   286: 'IGG_MESSAGE_WORD_02_BIT_5', class IGG Messages, trigger "64_Message_Data_IGG_MESSAGE_WORD_02" bit 13
   126: 'PIT-113 IGG MAIN ATOM AIR PRESSURE - FAULT', class BC Alarms, trigger "BC_ALARM_ACKNLG_4" bit 13
   125: 'TS-403 IG TEMP - HIGH HIGH SWITCH AND TIT-360 - FAULT', class BC Alarms, trigger "BC_ALARM_ACKNLG_4" bit 12
   128: 'TIT-202 IGG INLET FUEL TEMP', class BC Alarms, trigger "BC_ALARM_ACKNLG_4" bit 15
   127: 'PIT-205 IGG MAIN FUEL PRESSURE - FAULT', class BC Alarms, trigger "BC_ALARM_ACKNLG_4" bit 14
   313: 'BC_MESSAGE_WORD_02_BIT_0', class BC Messages, trigger "64_Message_Data_BC_MESSAGE_WORD_02" bit 8
   292: 'BC_MESSAGE_WORD_01_BIT_11', class BC Messages, trigger "64_Message_Data_BC_MESSAGE_WORD_01" bit 3
   311: 'BC_MESSAGE_WORD_02_BIT_14', class BC Messages, trigger "64_Message_Data_BC_MESSAGE_WORD_02" bit 6
   312: 'BC_MESSAGE_WORD_02_BIT_15', class BC Messages, trigger "64_Message_Data_BC_MESSAGE_WORD_02" bit 7
   289: 'BC_MESSAGE_WORD_01_BIT_8', class BC Messages, trigger "64_Message_Data_BC_MESSAGE_WORD_01" bit 0
   288: 'IGG_MESSAGE_WORD_02_BIT_7', class IGG Messages, trigger "64_Message_Data_IGG_MESSAGE_WORD_02" bit 15
   291: 'BC_MESSAGE_WORD_01_BIT_10', class BC Messages, trigger "64_Message_Data_BC_MESSAGE_WORD_01" bit 2
   290: 'BC_MESSAGE_WORD_01_BIT_9', class BC Messages, trigger "64_Message_Data_BC_MESSAGE_WORD_01" bit 1
   93: 'BC_ALARM_WORD_02_BIT_4', class BC Alarms, trigger "BC_ALARM_ACKNLG_2" bit 12
   75: 'BC AUTO INTERLOCKS NOT OK', class BC Alarms, trigger "BC_ALARM_ACKNLG_1" bit 10
   88: 'BC_ALARM_WORD_02_BIT_15', class BC Alarms, trigger "BC_ALARM_ACKNLG_2" bit 7
   283: 'IGG_MESSAGE_WORD_02_BIT_2', class IGG Messages, trigger "64_Message_Data_IGG_MESSAGE_WORD_02" bit 10
   320: 'BC_MESSAGE_WORD_02_BIT_7', class BC Messages, trigger "64_Message_Data_BC_MESSAGE_WORD_02" bit 15
   94: 'BC_ALARM_WORD_02_BIT_5', class BC Alarms, trigger "BC_ALARM_ACKNLG_2" bit 13
   74: 'IGNITER POWER NOT HEALTHY', class BC Alarms, trigger "BC_ALARM_ACKNLG_1" bit 9
   79: 'PILOT FLAME PURGE SEQUENCE FAILURE', class BC Alarms, trigger "BC_ALARM_ACKNLG_1" bit 14
   80: 'FD-001 FLAME DETECTION UNIT NOT HEALTHY', class BC Alarms, trigger "BC_ALARM_ACKNLG_1" bit 15
   84: 'PIT-204 FUEL OIL INLET PRESSURE LOW LOW AND PIT-205 - FAULT', class BC Alarms, trigger "BC_ALARM_ACKNLG_2" bit 3
   90: 'NO FLOW AT FS-320', class BC Alarms, trigger "BC_ALARM_ACKNLG_2" bit 9
   91: 'BC_ALARM_WORD_02_BIT_2', class BC Alarms, trigger "BC_ALARM_ACKNLG_2" bit 10
   83: 'BC_ALARM_WORD_02_BIT_10', class BC Alarms, trigger "BC_ALARM_ACKNLG_2" bit 2
   82: 'PIT-204 FUEL OIL INLET PRESSURE READING - FAULT AND CV-206 AND CV-207 - CLOSED', class BC Alarms, trigger "BC_ALARM_ACKNLG_2" bit 1
   76: 'FDU POWER NOT HEALTHY', class BC Alarms, trigger "BC_ALARM_ACKNLG_1" bit 11
   89: 'NO FLOW AT FS-317', class BC Alarms, trigger "BC_ALARM_ACKNLG_2" bit 8
   95: 'BC_ALARM_WORD_02_BIT_6', class BC Alarms, trigger "BC_ALARM_ACKNLG_2" bit 14
   87: 'PIT-204 FUEL OIL INLET PRESSURE - HIGH HIGH AND CV-206 AND CV-207 CLOSED', class BC Alarms, trigger "BC_ALARM_ACKNLG_2" bit 6
   85: 'PIT-204 FUEL OIL INLET PRESSURE - LOW LOW', class BC Alarms, trigger "BC_ALARM_ACKNLG_2" bit 4
   71: 'E-600 O2 ANALYSER CONTENT - LOW LOW', class BC Alarms, trigger "BC_ALARM_ACKNLG_1" bit 6
   77: 'PILOT FLAME IGNITION SEQUENCE FAILURE', class BC Alarms, trigger "BC_ALARM_ACKNLG_1" bit 12
   86: 'PIT-204 FUEL OIL INLET PRESSURE - HIGH HIGH AND PIT-205 - FAULT', class BC Alarms, trigger "BC_ALARM_ACKNLG_2" bit 5
   78: 'MAIN BURNER FLAME SEQUENCE FAILURE', class BC Alarms, trigger "BC_ALARM_ACKNLG_1" bit 13
   92: 'BC_ALARM_WORD_02_BIT_3', class BC Alarms, trigger "BC_ALARM_ACKNLG_2" bit 11
   96: 'BC_ALARM_WORD_02_BIT_7', class BC Alarms, trigger "BC_ALARM_ACKNLG_2" bit 15
   118: 'BC_ALARM_WORD_04_BIT_13', class BC Alarms, trigger "BC_ALARM_ACKNLG_4" bit 5
   72: 'E-600 O2 ANALYSER CONTENT - HIGH HIGH', class BC Alarms, trigger "BC_ALARM_ACKNLG_1" bit 7
   73: 'MASTER PLC HEART BEAT MISSING', class BC Alarms, trigger "BC_ALARM_ACKNLG_1" bit 8
   81: 'PIT-204 FUEL OIL INLET PRESSURE READING - FAULT AND PIT-205 - FAULT', class BC Alarms, trigger "BC_ALARM_ACKNLG_2" bit 0
   319: 'BC_MESSAGE_WORD_02_BIT_6', class BC Messages, trigger "64_Message_Data_BC_MESSAGE_WORD_02" bit 14
   385: 'IGG_WARNING_WORD_01_BIT_8', class IGG Warnings, trigger "62_Warning_Data_IGG_WARNING_WORD_01" bit 0
   386: 'IGG_WARNING_WORD_01_BIT_9', class IGG Warnings, trigger "62_Warning_Data_IGG_WARNING_WORD_01" bit 1
   387: 'IGG_WARNING_WORD_01_BIT_10', class IGG Warnings, trigger "62_Warning_Data_IGG_WARNING_WORD_01" bit 2
   388: 'IGG_WARNING_WORD_01_BIT_11', class IGG Warnings, trigger "62_Warning_Data_IGG_WARNING_WORD_01" bit 3
   389: 'IGG_WARNING_WORD_01_BIT_12', class IGG Warnings, trigger "62_Warning_Data_IGG_WARNING_WORD_01" bit 4
   390: 'IGG_WARNING_WORD_01_BIT_13', class IGG Warnings, trigger "62_Warning_Data_IGG_WARNING_WORD_01" bit 5
   391: 'IGG_WARNING_WORD_01_BIT_14', class IGG Warnings, trigger "62_Warning_Data_IGG_WARNING_WORD_01" bit 6
   392: 'IGG_WARNING_WORD_01_BIT_15', class IGG Warnings, trigger "62_Warning_Data_IGG_WARNING_WORD_01" bit 7
   393: '31B1 ATMOSPHERIC O2 SENSOR - LOW', class IGG Warnings, trigger "62_Warning_Data_IGG_WARNING_WORD_01" bit 8
   394: '31B2 ATMOSPHERIC O2 SENSOR - LOW', class IGG Warnings, trigger "62_Warning_Data_IGG_WARNING_WORD_01" bit 9
   395: '31B1 ATMOSPHERIC O2 SENSOR - LOW LOW', class IGG Warnings, trigger "62_Warning_Data_IGG_WARNING_WORD_01" bit 10
   396: '31B2 ATMOSPHERIC O2 SENSOR - LOW LOW', class IGG Warnings, trigger "62_Warning_Data_IGG_WARNING_WORD_01" bit 11
   397: 'IGG_WARNING_WORD_01_BIT_4', class IGG Warnings, trigger "62_Warning_Data_IGG_WARNING_WORD_01" bit 12
   398: 'IGG_WARNING_WORD_01_BIT_5', class IGG Warnings, trigger "62_Warning_Data_IGG_WARNING_WORD_01" bit 13
   399: 'IGG_WARNING_WORD_01_BIT_6', class IGG Warnings, trigger "62_Warning_Data_IGG_WARNING_WORD_01" bit 14
   400: 'IGG_WARNING_WORD_01_BIT_7', class IGG Warnings, trigger "62_Warning_Data_IGG_WARNING_WORD_01" bit 15
   401: 'PIT-359 INLET CSW PRESSURE - LOW', class IGG Warnings, trigger "62_Warning_Data_IGG_WARNING_WORD_02" bit 0
   402: 'PIT-359 INLET CSW PRESSURE - HIGH', class IGG Warnings, trigger "62_Warning_Data_IGG_WARNING_WORD_02" bit 1
   403: 'PIT-316 OUTLET CSW PRESSURE - LOW', class IGG Warnings, trigger "62_Warning_Data_IGG_WARNING_WORD_02" bit 2
   404: 'PIT-316 OUTLET CSW PRESSURE - HIGH', class IGG Warnings, trigger "62_Warning_Data_IGG_WARNING_WORD_02" bit 3
   405: 'PIT-316 OUTLET CSW PRESSURE - LOW LOW', class IGG Warnings, trigger "62_Warning_Data_IGG_WARNING_WORD_02" bit 4
   406: 'PIT-316 OUTLET CSW PRESSURE - HIGH HIGH', class IGG Warnings, trigger "62_Warning_Data_IGG_WARNING_WORD_02" bit 5
   407: 'IGG_WARNING_WORD_02_BIT_14', class IGG Warnings, trigger "62_Warning_Data_IGG_WARNING_WORD_02" bit 6
   408: 'IGG_WARNING_WORD_02_BIT_15', class IGG Warnings, trigger "62_Warning_Data_IGG_WARNING_WORD_02" bit 7
   409: 'PIT-102 CA PRESSURE LOW', class IGG Warnings, trigger "62_Warning_Data_IGG_WARNING_WORD_02" bit 8
   410: 'PIT-102 CA PRESSURE HIGH', class IGG Warnings, trigger "62_Warning_Data_IGG_WARNING_WORD_02" bit 9
   411: 'TIT-401 IG TEMP HIGH', class IGG Warnings, trigger "62_Warning_Data_IGG_WARNING_WORD_02" bit 10
   412: 'PIT-402 IG OUTLET PRESSURE - LOW', class IGG Warnings, trigger "62_Warning_Data_IGG_WARNING_WORD_02" bit 11
   413: 'PIT-402 IG OUTLET PRESSURE - HIGH', class IGG Warnings, trigger "62_Warning_Data_IGG_WARNING_WORD_02" bit 12
   414: 'TIT-315 SHELL CSW TEMP - HIGH', class IGG Warnings, trigger "62_Warning_Data_IGG_WARNING_WORD_02" bit 13
   415: 'TIT-319 INLET CSW TEMP - HIGH', class IGG Warnings, trigger "62_Warning_Data_IGG_WARNING_WORD_02" bit 14
   416: 'TIT-360 OUTLET CSW TEMP - HIGH', class IGG Warnings, trigger "62_Warning_Data_IGG_WARNING_WORD_02" bit 15
   417: 'FD-001 FLAME - TRIPPED', class BC Warnings, trigger "62_Warning_Data_BC_WARNING_WORD_01" bit 0
   418: 'PIT-204 FUEL OIL INLET PRESSURE - LOW LOW', class BC Warnings, trigger "62_Warning_Data_BC_WARNING_WORD_01" bit 1
   419: 'PIT-204 FUEL OIL INLET PRESSURE - LOW', class BC Warnings, trigger "62_Warning_Data_BC_WARNING_WORD_01" bit 2
   420: 'PIT-204 FUEL OIL INLET PRESSURE - HIGH', class BC Warnings, trigger "62_Warning_Data_BC_WARNING_WORD_01" bit 3
   421: 'PIT-204 FUEL OIL INLET PRESSURE - HIGH HIGH', class BC Warnings, trigger "62_Warning_Data_BC_WARNING_WORD_01" bit 4
   422: 'PIT-204 FUEL OIL INLET PRESSURE - OUT OF RANGE', class BC Warnings, trigger "62_Warning_Data_BC_WARNING_WORD_01" bit 5
   423: 'BC_WARNING_WORD_01_BIT_14', class BC Warnings, trigger "62_Warning_Data_BC_WARNING_WORD_01" bit 6
   424: 'BC_WARNING_WORD_01_BIT_15', class BC Warnings, trigger "62_Warning_Data_BC_WARNING_WORD_01" bit 7
   425: 'BC_WARNING_WORD_01_BIT_0', class BC Warnings, trigger "62_Warning_Data_BC_WARNING_WORD_01" bit 8
   426: 'PIT-204 FUEL OIL INLET PRESSURE - LOW LOW', class BC Warnings, trigger "62_Warning_Data_BC_WARNING_WORD_01" bit 9
   427: 'PIT-204 FUEL OIL INLET PRESSURE - LOW', class BC Warnings, trigger "62_Warning_Data_BC_WARNING_WORD_01" bit 10
   428: 'PIT-204 FUEL OIL INLET PRESSURE - HIGH', class BC Warnings, trigger "62_Warning_Data_BC_WARNING_WORD_01" bit 11
   429: 'PIT-204 FUEL OIL INLET PRESSURE - HIGH HIGH', class BC Warnings, trigger "62_Warning_Data_BC_WARNING_WORD_01" bit 12
   430: 'PIT-204 FUEL OIL INLET PRESSURE - OUT OF RANGE', class BC Warnings, trigger "62_Warning_Data_BC_WARNING_WORD_01" bit 13
   431: 'FD-001 FLAME NOT DETECTED', class BC Warnings, trigger "62_Warning_Data_BC_WARNING_WORD_01" bit 14
   432: 'FD-001 FLAME NOT HEALTHY', class BC Warnings, trigger "62_Warning_Data_BC_WARNING_WORD_01" bit 15
   433: 'BC_WARNING_WORD_02_BIT_8', class BC Warnings, trigger "62_Warning_Data_BC_WARNING_WORD_02" bit 0
   434: 'TIT-202 FUEL OIL INLET TEMPERATURE - LOW LOW', class BC Warnings, trigger "62_Warning_Data_BC_WARNING_WORD_02" bit 1
   435: 'TIT-202 FUEL OIL INLET TEMPERATURE - LOW', class BC Warnings, trigger "62_Warning_Data_BC_WARNING_WORD_02" bit 2
   436: 'TIT-202 FUEL OIL INLET TEMPERATURE - HIGH', class BC Warnings, trigger "62_Warning_Data_BC_WARNING_WORD_02" bit 3
   437: 'TIT-202 FUEL OIL INLET TEMPERATURE - HIGH HIGH', class BC Warnings, trigger "62_Warning_Data_BC_WARNING_WORD_02" bit 4
   438: 'TIT-202 FUEL OIL INLET TEMPERATURE - OUT OF RANGE', class BC Warnings, trigger "62_Warning_Data_BC_WARNING_WORD_02" bit 5
   439: 'BC_WARNING_WORD_02_BIT_14', class BC Warnings, trigger "62_Warning_Data_BC_WARNING_WORD_02" bit 6
   440: 'BC_WARNING_WORD_02_BIT_15', class BC Warnings, trigger "62_Warning_Data_BC_WARNING_WORD_02" bit 7
   441: 'BC_WARNING_WORD_02_BIT_0', class BC Warnings, trigger "62_Warning_Data_BC_WARNING_WORD_02" bit 8
   442: 'TIT-202 IGG INLET FUEL TEMP - LOW LOW', class BC Warnings, trigger "62_Warning_Data_BC_WARNING_WORD_02" bit 9
   443: 'TIT-202 IGG INLET FUEL TEMP - LOW', class BC Warnings, trigger "62_Warning_Data_BC_WARNING_WORD_02" bit 10
   444: 'TIT-202 IGG INLET FUEL TEMP - HIGH', class BC Warnings, trigger "62_Warning_Data_BC_WARNING_WORD_02" bit 11
   445: 'TIT-202 IGG INLET FUEL TEMP - HIGH HIGH', class BC Warnings, trigger "62_Warning_Data_BC_WARNING_WORD_02" bit 12
   446: 'TIT-202 IGG INLET FUEL TEMP - OUT OF RANGE', class BC Warnings, trigger "62_Warning_Data_BC_WARNING_WORD_02" bit 13
   447: 'BC_WARNING_WORD_02_BIT_6', class BC Warnings, trigger "62_Warning_Data_BC_WARNING_WORD_02" bit 14
   448: 'BC_WARNING_WORD_02_BIT_7', class BC Warnings, trigger "62_Warning_Data_BC_WARNING_WORD_02" bit 15
   449: 'PIT-102 CA PRESSURE - LOW LOW', class IGG Warnings, trigger "62_Warning_Data_IGG_WARNING_WORD_03" bit 0
   450: 'PIT-102 CA PRESSURE - HIGH HIGH', class IGG Warnings, trigger "62_Warning_Data_IGG_WARNING_WORD_03" bit 1
   451: 'IGG WARNING', class IGG Warnings, trigger "62_Warning_Data_IGG_WARNING_WORD_03" bit 2
   452: 'PIT-402 IG OUTLET PRESSURE - LOW LOW', class IGG Warnings, trigger "62_Warning_Data_IGG_WARNING_WORD_03" bit 3
   453: 'PIT-402 IG OUTLET PRESSURE - HIGH HIGH', class IGG Warnings, trigger "62_Warning_Data_IGG_WARNING_WORD_03" bit 4
   454: 'TIT-315 SHELL CSW TEMP - HIGH HIGH', class IGG Warnings, trigger "62_Warning_Data_IGG_WARNING_WORD_03" bit 5
   455: 'TIT-319 INLET CSW TEMP - HIGH HIGH', class IGG Warnings, trigger "62_Warning_Data_IGG_WARNING_WORD_03" bit 6
   456: 'TIT-360 OUTLET CSW TEMP - HIGH HIGH', class IGG Warnings, trigger "62_Warning_Data_IGG_WARNING_WORD_03" bit 7
   457: 'PIT-112 IA PRESSURE- OUT OF RANGE', class IGG Warnings, trigger "62_Warning_Data_IGG_WARNING_WORD_03" bit 8
   458: 'PIT-113 FUEL PRESSURE TO MAIN BURNER - OUT OF RANGE', class IGG Warnings, trigger "62_Warning_Data_IGG_WARNING_WORD_03" bit 9
   459: 'PIT-102 CA PRESSURE - OUT OF RANGE', class IGG Warnings, trigger "62_Warning_Data_IGG_WARNING_WORD_03" bit 10
   460: 'TIT-401 IG TEMP - OUT OF RANGE', class IGG Warnings, trigger "62_Warning_Data_IGG_WARNING_WORD_03" bit 11
   461: 'PIT-402 IG VENT PRESSURE - OUT OF RANGE', class IGG Warnings, trigger "62_Warning_Data_IGG_WARNING_WORD_03" bit 12
   462: 'TIT-315 SHELL CSW TEMP - OUT OF RANGE', class IGG Warnings, trigger "62_Warning_Data_IGG_WARNING_WORD_03" bit 13
   463: 'TIT-319 INLET CSW TEMP - OUT OF RANGE', class IGG Warnings, trigger "62_Warning_Data_IGG_WARNING_WORD_03" bit 14
   464: 'TIT-360 OUTLET CSW TEMP - OUT OF RANGE', class IGG Warnings, trigger "62_Warning_Data_IGG_WARNING_WORD_03" bit 15
   465: 'INTERLOCKS NOT OK', class IGG Warnings, trigger "62_Warning_Data_IGG_WARNING_WORD_04" bit 0
   466: 'CHECK PIT-316 - WARNING', class IGG Warnings, trigger "62_Warning_Data_IGG_WARNING_WORD_04" bit 1
   467: 'CHECK PIT-102 - WARNING', class IGG Warnings, trigger "62_Warning_Data_IGG_WARNING_WORD_04" bit 2
   468: 'CHECK PIT-102 - WARNING II', class IGG Warnings, trigger "62_Warning_Data_IGG_WARNING_WORD_04" bit 3
   469: 'CHECK TIT-401 - WARNING', class IGG Warnings, trigger "62_Warning_Data_IGG_WARNING_WORD_04" bit 4
   470: 'CHECK TIT-319 - WARNING', class IGG Warnings, trigger "62_Warning_Data_IGG_WARNING_WORD_04" bit 5
   471: 'CHECK TIT-360 - WARNING', class IGG Warnings, trigger "62_Warning_Data_IGG_WARNING_WORD_04" bit 6
   472: 'E-500A TRIPPED', class IGG Warnings, trigger "62_Warning_Data_IGG_WARNING_WORD_04" bit 7
   473: 'E-500B TRIPPED', class IGG Warnings, trigger "62_Warning_Data_IGG_WARNING_WORD_04" bit 8
   474: 'PIT-359 INLET CSW PRESSURE - LOW LOW', class IGG Warnings, trigger "62_Warning_Data_IGG_WARNING_WORD_04" bit 9
   475: 'PIT-359 INLET CSW PRESSURE - HIGH HIGH', class IGG Warnings, trigger "62_Warning_Data_IGG_WARNING_WORD_04" bit 10
   476: 'PIT-359 INLET CSW PRESSURE - OUT OF RANGE', class IGG Warnings, trigger "62_Warning_Data_IGG_WARNING_WORD_04" bit 11
   477: 'PIT-316 OUTLET CSW PRESSURE - OUT OF RANGE', class IGG Warnings, trigger "62_Warning_Data_IGG_WARNING_WORD_04" bit 12
   478: 'PIT-112 IA PRESSURE - OUT OF RANGE', class IGG Warnings, trigger "62_Warning_Data_IGG_WARNING_WORD_04" bit 13
   479: 'IGG_WARNING_WORD_04_BIT_6', class IGG Warnings, trigger "62_Warning_Data_IGG_WARNING_WORD_04" bit 14
   480: 'IGG_WARNING_WORD_04_BIT_7', class IGG Warnings, trigger "62_Warning_Data_IGG_WARNING_WORD_04" bit 15
   481: 'BC_WARNING_WORD_03_BIT_8', class BC Warnings, trigger "62_Warning_Data_BC_WARNING_WORD_03" bit 0
   482: 'E-600 O2 ANALYSER CONTENT HIGH HIGH', class BC Warnings, trigger "62_Warning_Data_BC_WARNING_WORD_03" bit 1
   483: 'BC_WARNING_WORD_03_BIT_10', class BC Warnings, trigger "62_Warning_Data_BC_WARNING_WORD_03" bit 2
   484: 'BC_WARNING_WORD_03_BIT_11', class BC Warnings, trigger "62_Warning_Data_BC_WARNING_WORD_03" bit 3
   485: 'BC_WARNING_WORD_03_BIT_12', class BC Warnings, trigger "62_Warning_Data_BC_WARNING_WORD_03" bit 4
   486: 'BC_WARNING_WORD_03_BIT_13', class BC Warnings, trigger "62_Warning_Data_BC_WARNING_WORD_03" bit 5
   487: 'IGNITER POWER - NOT HEALTHY', class BC Warnings, trigger "62_Warning_Data_BC_WARNING_WORD_03" bit 6
   488: 'BC_WARNING_WORD_03_BIT_13', class BC Warnings, trigger "62_Warning_Data_BC_WARNING_WORD_03" bit 7
   489: 'BC_WARNING_WORD_03_BIT_0', class BC Warnings, trigger "62_Warning_Data_BC_WARNING_WORD_03" bit 8
   490: 'PIT-205 IGG MAIN FUEL PRESSURE - LOW', class BC Warnings, trigger "62_Warning_Data_BC_WARNING_WORD_03" bit 9
   491: 'PIT-205 IGG MAIN FUEL PRESSURE - LOW LOW', class BC Warnings, trigger "62_Warning_Data_BC_WARNING_WORD_03" bit 10
   492: 'PIT-205 IGG MAIN FUEL PRESSURE - HIGH', class BC Warnings, trigger "62_Warning_Data_BC_WARNING_WORD_03" bit 11
   493: 'PIT-205 IGG MAIN FUEL PRESSURE - HIGH HIGH', class BC Warnings, trigger "62_Warning_Data_BC_WARNING_WORD_03" bit 12
   494: 'PIT-205 IGG MAIN FUEL PRESSURE - OUT OF RANGE', class BC Warnings, trigger "62_Warning_Data_BC_WARNING_WORD_03" bit 13
   495: 'E-131 IA COMPRESSOR - WARNING', class BC Warnings, trigger "62_Warning_Data_BC_WARNING_WORD_03" bit 14
   496: 'E-131 IA COMPRESSOR - NOT RUNNING', class BC Warnings, trigger "62_Warning_Data_BC_WARNING_WORD_03" bit 15
   497: 'CHECK PIT-112 IA PRESSURE - WARNING', class BC Warnings, trigger "62_Warning_Data_BC_WARNING_WORD_04" bit 0
   498: 'CHECK PIT-204 FUEL OIL INLET PRESSURE - WARNING', class BC Warnings, trigger "62_Warning_Data_BC_WARNING_WORD_04" bit 1
   499: 'CHECK FS-123 PILOT AIR FLOW - WARNING', class BC Warnings, trigger "62_Warning_Data_BC_WARNING_WORD_04" bit 2
   500: 'CHECK FS-115 MAIN BURNER ATOMISING AIR FLOW - WARNING', class BC Warnings, trigger "62_Warning_Data_BC_WARNING_WORD_04" bit 3
   501: 'CHECK FS-317 IGG JACKET COOLING WATER FLOW - WARNING', class BC Warnings, trigger "62_Warning_Data_BC_WARNING_WORD_04" bit 4
   502: 'SOOT SYSTEM POWER - NOT HEALTHY', class BC Warnings, trigger "62_Warning_Data_BC_WARNING_WORD_04" bit 5
   503: 'SOOT SYSTEM OPACITY - HIGH', class BC Warnings, trigger "62_Warning_Data_BC_WARNING_WORD_04" bit 6
   504: 'SOOT SYSTEM - OUT OF RANGE', class BC Warnings, trigger "62_Warning_Data_BC_WARNING_WORD_04" bit 7
   505: 'BC_INTERLOCKS NOT OK', class BC Warnings, trigger "62_Warning_Data_BC_WARNING_WORD_04" bit 8
   506: 'PIT-112 INLET IA PRESSURE - LOW LOW', class BC Warnings, trigger "62_Warning_Data_BC_WARNING_WORD_04" bit 9
   507: 'PIT-112 INLET IA PRESSURE - LOW', class BC Warnings, trigger "62_Warning_Data_BC_WARNING_WORD_04" bit 10
   508: 'PIT-112 INLET IA PRESSURE - HIGH', class BC Warnings, trigger "62_Warning_Data_BC_WARNING_WORD_04" bit 11
   509: 'PIT-112 INLET IA PRESSURE - HIGH HIGH', class BC Warnings, trigger "62_Warning_Data_BC_WARNING_WORD_04" bit 12
   510: 'PIT-112 INLET IA PRESSURE - OUT OF RANGE', class BC Warnings, trigger "62_Warning_Data_BC_WARNING_WORD_04" bit 13
   511: 'CHECK FS-317 IGG JACKET COOLING WATER FLOW - WARNING', class BC Warnings, trigger "62_Warning_Data_BC_WARNING_WORD_04" bit 14
   512: 'CHECK FS-320 REAR MATRIX COOLING WATER FLOW - WARNING', class BC Warnings, trigger "62_Warning_Data_BC_WARNING_WORD_04" bit 15
   513: 'IGG HMI LOST COMUNICATION', class IGG Warnings, trigger "62_Warning_Data_IGG_WARNING_WORD_05" bit 0
   514: 'CCR HMI LOST COMUNICATION', class IGG Warnings, trigger "62_Warning_Data_IGG_WARNING_WORD_05" bit 1
   515: 'BRIGE HMI LOST COMUNICATION', class IGG Warnings, trigger "62_Warning_Data_IGG_WARNING_WORD_05" bit 2
   516: 'PIT-402 CA PRESSURE - LOW LOW', class IGG Warnings, trigger "62_Warning_Data_IGG_WARNING_WORD_05" bit 3
   517: 'PIT-402 CA PRESSURE - HIGH HIGH', class IGG Warnings, trigger "62_Warning_Data_IGG_WARNING_WORD_05" bit 4
   518: 'TIT-315 SHELL CSW TEMP - HIGH HIGH', class IGG Warnings, trigger "62_Warning_Data_IGG_WARNING_WORD_05" bit 5
   519: 'TIT-319 INLET CSW TEMP - HIGH HIGH', class IGG Warnings, trigger "62_Warning_Data_IGG_WARNING_WORD_05" bit 6
   520: 'TIT-360 OUTLET CSW TEMP - HIGH HIGH', class IGG Warnings, trigger "62_Warning_Data_IGG_WARNING_WORD_05" bit 7
   521: 'BC PLC POWER NOT HEALTHY', class IGG Warnings, trigger "62_Warning_Data_IGG_WARNING_WORD_05" bit 8
   522: 'CONTROLS POWER SUPPLY - NOT HEALTHY', class IGG Warnings, trigger "62_Warning_Data_IGG_WARNING_WORD_05" bit 9
   523: 'IGG POWER SUPPLY - NOT HEALTHY', class IGG Warnings, trigger "62_Warning_Data_IGG_WARNING_WORD_05" bit 10
   524: 'BC POWER SUPPLY - NOT HEALTHY', class IGG Warnings, trigger "62_Warning_Data_IGG_WARNING_WORD_05" bit 11
   525: 'BACKUP 24VDC POWER SUPPLY - NOT HEALTHY', class IGG Warnings, trigger "62_Warning_Data_IGG_WARNING_WORD_05" bit 12
   526: 'IGG VENTILATION POWER - NOT HEALTHY', class IGG Warnings, trigger "62_Warning_Data_IGG_WARNING_WORD_05" bit 13
   527: 'MCCP VENTILATION POWER - NOT HEALTHY', class IGG Warnings, trigger "62_Warning_Data_IGG_WARNING_WORD_05" bit 14
   528: 'TIT-360 OUTLET CSW TEMP - HIGH HIGH', class IGG Warnings, trigger "62_Warning_Data_IGG_WARNING_WORD_05" bit 15
   529: 'PIT-359 INLET CSW PRESSURE - LOW LOW', class IGG Warnings, trigger "62_Warning_Data_IGG_WARNING_WORD_06" bit 0
   530: 'PIT-359 INLET CSW PRESSURE - HIGH HIGH', class IGG Warnings, trigger "62_Warning_Data_IGG_WARNING_WORD_06" bit 1
   531: 'IGG_WARNING_WORD_06_BIT_10', class IGG Warnings, trigger "62_Warning_Data_IGG_WARNING_WORD_06" bit 2
   532: 'IGG_WARNING_WORD_06_BIT_11', class IGG Warnings, trigger "62_Warning_Data_IGG_WARNING_WORD_06" bit 3
   533: 'IGG_WARNING_WORD_06_BIT_12', class IGG Warnings, trigger "62_Warning_Data_IGG_WARNING_WORD_06" bit 4
   534: 'IGG_WARNING_WORD_06_BIT_13', class IGG Warnings, trigger "62_Warning_Data_IGG_WARNING_WORD_06" bit 5
   535: 'IGG_WARNING_WORD_06_BIT_14', class IGG Warnings, trigger "62_Warning_Data_IGG_WARNING_WORD_06" bit 6
   536: 'IGG_WARNING_WORD_06_BIT_15', class IGG Warnings, trigger "62_Warning_Data_IGG_WARNING_WORD_06" bit 7
   537: 'IGG_WARNING_WORD_06_BIT_0', class IGG Warnings, trigger "62_Warning_Data_IGG_WARNING_WORD_06" bit 8
   538: 'IGG_WARNING_WORD_06_BIT_1', class IGG Warnings, trigger "62_Warning_Data_IGG_WARNING_WORD_06" bit 9
   539: 'IGG_WARNING_WORD_06_BIT_2', class IGG Warnings, trigger "62_Warning_Data_IGG_WARNING_WORD_06" bit 10
   540: 'IGG_WARNING_WORD_06_BIT_3', class IGG Warnings, trigger "62_Warning_Data_IGG_WARNING_WORD_06" bit 11
   541: 'IGG_WARNING_WORD_06_BIT_4', class IGG Warnings, trigger "62_Warning_Data_IGG_WARNING_WORD_06" bit 12
   542: 'IGG_WARNING_WORD_06_BIT_5', class IGG Warnings, trigger "62_Warning_Data_IGG_WARNING_WORD_06" bit 13
   543: 'IGG_WARNING_WORD_06_BIT_6', class IGG Warnings, trigger "62_Warning_Data_IGG_WARNING_WORD_06" bit 14
   544: 'IGG_WARNING_WORD_06_BIT_7', class IGG Warnings, trigger "62_Warning_Data_IGG_WARNING_WORD_06" bit 15
   545: 'BC_WARNING_WORD_05_BIT_8', class BC Warnings, trigger "62_Warning_Data_BC_WARNING_WORD_05" bit 0
   546: 'BC_WARNING_WORD_05_BIT_9', class BC Warnings, trigger "62_Warning_Data_BC_WARNING_WORD_05" bit 1
   547: 'BC_WARNING_WORD_05_BIT_10', class BC Warnings, trigger "62_Warning_Data_BC_WARNING_WORD_05" bit 2
   548: 'BC_WARNING_WORD_05_BIT_11', class BC Warnings, trigger "62_Warning_Data_BC_WARNING_WORD_05" bit 3
   549: 'BC_WARNING_WORD_05_BIT_12', class BC Warnings, trigger "62_Warning_Data_BC_WARNING_WORD_05" bit 4
   550: 'BC_WARNING_WORD_05_BIT_13', class BC Warnings, trigger "62_Warning_Data_BC_WARNING_WORD_05" bit 5
   551: 'BC_WARNING_WORD_05_BIT_14', class BC Warnings, trigger "62_Warning_Data_BC_WARNING_WORD_05" bit 6
   552: 'BC_WARNING_WORD_05_BIT_15', class BC Warnings, trigger "62_Warning_Data_BC_WARNING_WORD_05" bit 7
   553: 'BC_WARNING_WORD_05_BIT_0', class BC Warnings, trigger "62_Warning_Data_BC_WARNING_WORD_05" bit 8
   554: 'PIT-113 IGG MAIN ATOM AIR PRESSURE - LOW LOW', class BC Warnings, trigger "62_Warning_Data_BC_WARNING_WORD_05" bit 9
   555: 'PIT-113 IGG MAIN ATOM AIR PRESSURE - LOW', class BC Warnings, trigger "62_Warning_Data_BC_WARNING_WORD_05" bit 10
   556: 'PIT-113 IGG MAIN ATOM AIR PRESSURE - HIGH', class BC Warnings, trigger "62_Warning_Data_BC_WARNING_WORD_05" bit 11
   557: 'PIT-113 IGG MAIN ATOM AIR PRESSURE - HIGH HIGH', class BC Warnings, trigger "62_Warning_Data_BC_WARNING_WORD_05" bit 12
   558: 'PIT-113 IGG MAIN ATOM AIR PRESSURE - OUT OF RANGE', class BC Warnings, trigger "62_Warning_Data_BC_WARNING_WORD_05" bit 13
   559: 'BC_WARNING_WORD', class BC Warnings, trigger "62_Warning_Data_BC_WARNING_WORD_05" bit 14
   560: 'BC_WARNING WORD', class BC Warnings, trigger "62_Warning_Data_BC_WARNING_WORD_05" bit 15
   561: 'INTERLOCKS NOT OK', class BC Warnings, trigger "62_Warning_Data_BC_WARNING_WORD_06" bit 0
   562: 'BC_WARNING_WORD_06_BIT_9', class BC Warnings, trigger "62_Warning_Data_BC_WARNING_WORD_06" bit 1
   563: 'BC_WARNING_WORD_06_BIT_10', class BC Warnings, trigger "62_Warning_Data_BC_WARNING_WORD_06" bit 2
   564: 'BC_WARNING_WORD_06_BIT_11', class BC Warnings, trigger "62_Warning_Data_BC_WARNING_WORD_06" bit 3
   565: 'BC_WARNING_WORD_06_BIT_12', class BC Warnings, trigger "62_Warning_Data_BC_WARNING_WORD_06" bit 4
   566: 'BC_WARNING_WORD_06_BIT_13', class BC Warnings, trigger "62_Warning_Data_BC_WARNING_WORD_06" bit 5
   567: 'BC_WARNING_WORD_06_BIT_14', class BC Warnings, trigger "62_Warning_Data_BC_WARNING_WORD_06" bit 6
   568: 'BC_WARNING_WORD_06_BIT_15', class BC Warnings, trigger "62_Warning_Data_BC_WARNING_WORD_06" bit 7
   569: 'INTERLOCKS NOT OK', class BC Warnings, trigger "62_Warning_Data_BC_WARNING_WORD_06" bit 8
   570: 'BC_WARNING_WORD_06_BIT_1', class BC Warnings, trigger "62_Warning_Data_BC_WARNING_WORD_06" bit 9
   571: 'BC_WARNING_WORD_06_BIT_2', class BC Warnings, trigger "62_Warning_Data_BC_WARNING_WORD_06" bit 10
   572: 'BC_WARNING_WORD_06_BIT_3', class BC Warnings, trigger "62_Warning_Data_BC_WARNING_WORD_06" bit 11
   573: 'BC_WARNING_WORD_06_BIT_4', class BC Warnings, trigger "62_Warning_Data_BC_WARNING_WORD_06" bit 12
   574: 'BC_WARNING_WORD_06_BIT_5', class BC Warnings, trigger "62_Warning_Data_BC_WARNING_WORD_06" bit 13
   575: 'BC_WARNING_WORD_06_BIT_6', class BC Warnings, trigger "62_Warning_Data_BC_WARNING_WORD_06" bit 14
   576: 'BC_WARNING_WORD_06_BIT_7', class BC Warnings, trigger "62_Warning_Data_BC_WARNING_WORD_06" bit 15
   577: 'BC_WARNING_WORD_05_BIT_8', class BC Warnings bit 0
   2182: 'FIT418 7 APT TANK USD FLOW LOW', class Tank Control Warnings, trigger "2062_Warning_Data_BTCS_WARNING_WORD_04" bit 6
   2183: 'FIT418 7 APT TANK USD FLOW HIGH', class Tank Control Warnings, trigger "2062_Warning_Data_BTCS_WARNING_WORD_04" bit 7
   2181: 'FIT417 6 STARBOARD TANK USD FLOW HIGH', class Tank Control Warnings, trigger "2062_Warning_Data_BTCS_WARNING_WORD_04" bit 5
   2179: 'FIT418 6 PORT TANK USD FLOW HIGH', class Tank Control Warnings, trigger "2062_Warning_Data_BTCS_WARNING_WORD_04" bit 3
   2180: 'FIT417 6 STARBOARD TANK USD FLOW LOW', class Tank Control Warnings, trigger "2062_Warning_Data_BTCS_WARNING_WORD_04" bit 4
   2184: 'FIT417 3 STARBOARD TANK USD FLOW LOW', class Tank Control Warnings, trigger "2062_Warning_Data_BTCS_WARNING_WORD_04" bit 8
   2275: 'LT422 5 PORT TANK LEVEL LOW', class Tank Control Warnings, trigger "2062_Warning_Data_BTCS_WARNING_WORD_10" bit 3
   2185: 'FIT417 3 STARBOARD TANK USD FLOW HIGH', class Tank Control Warnings, trigger "2062_Warning_Data_BTCS_WARNING_WORD_04" bit 9
   2274: 'LT422 5 PORT TANK LEVEL HIGH', class Tank Control Warnings, trigger "2062_Warning_Data_BTCS_WARNING_WORD_10" bit 2
   2272: 'LT422 4 STARBOARD TANK LEVEL HIGH', class Tank Control Warnings, trigger "2062_Warning_Data_BTCS_WARNING_WORD_10" bit 0
   2273: 'LT422 4 STARBOARD TANK LEVEL LOW', class Tank Control Warnings, trigger "2062_Warning_Data_BTCS_WARNING_WORD_10" bit 1
   2171: 'TT-426 7 AFT PEACK TANK TEMPERATURE - HIGH', class Tank Control Warnings, trigger "2062_Warning_Data_BTCS_WARNING_WORD_03" bit 11
   2172: 'BTCS_WARNING_WORD_03_BIT_4', class Tank Control Warnings, trigger "2062_Warning_Data_BTCS_WARNING_WORD_03" bit 12
   2170: 'TT-426 6 STARBOARD TANK TEMPERATURE - HIGH', class Tank Control Warnings, trigger "2062_Warning_Data_BTCS_WARNING_WORD_03" bit 10
   2168: 'TT-426 5 STARBOARD TANK TEMPERATURE - HIGH', class Tank Control Warnings, trigger "2062_Warning_Data_BTCS_WARNING_WORD_03" bit 8
   2169: 'TT-426 6 PORT TANK TEMPERATURE - HIGH', class Tank Control Warnings, trigger "2062_Warning_Data_BTCS_WARNING_WORD_03" bit 9
   2173: 'BTCS_WARNING_WORD_03_BIT_5', class Tank Control Warnings, trigger "2062_Warning_Data_BTCS_WARNING_WORD_03" bit 13
   2177: 'FIT417 5 STARBOARD TANK USD FLOW HIGH', class Tank Control Warnings, trigger "2062_Warning_Data_BTCS_WARNING_WORD_04" bit 1
   2178: 'FIT418 6 PORT TANK USD FLOW LOW', class Tank Control Warnings, trigger "2062_Warning_Data_BTCS_WARNING_WORD_04" bit 2
   2176: 'FIT417 5 STARBOARD TANK USD FLOW LOW', class Tank Control Warnings, trigger "2062_Warning_Data_BTCS_WARNING_WORD_04" bit 0
   2174: 'BTCS_WARNING_WORD_03_BIT_6', class Tank Control Warnings, trigger "2062_Warning_Data_BTCS_WARNING_WORD_03" bit 14
   2175: 'BTCS_WARNING_WORD_03_BIT_7', class Tank Control Warnings, trigger "2062_Warning_Data_BTCS_WARNING_WORD_03" bit 15
   2186: 'FIT418 4 PORT TANK USD FLOW LOW', class Tank Control Warnings, trigger "2062_Warning_Data_BTCS_WARNING_WORD_04" bit 10
   2195: 'FIT420 4 PORT MBG FLOW HIGH', class Tank Control Warnings, trigger "2062_Warning_Data_BTCS_WARNING_WORD_05" bit 3
   2282: 'LT422 3 PORT TANK LEVEL HIGH', class Tank Control Warnings, trigger "2062_Warning_Data_BTCS_WARNING_WORD_10" bit 10
   2281: 'LT422 2 STARBOARD TANK LEVEL LOW', class Tank Control Warnings, trigger "2062_Warning_Data_BTCS_WARNING_WORD_10" bit 9
   2193: 'FIT419 3 STARBOARD MBG FLOW HIGH', class Tank Control Warnings, trigger "2062_Warning_Data_BTCS_WARNING_WORD_05" bit 1
   2194: 'FIT420 4 PORT MBG FLOW LOW', class Tank Control Warnings, trigger "2062_Warning_Data_BTCS_WARNING_WORD_05" bit 2
   2196: 'FIT419 4 STARBOARD MBG FLOW LOW', class Tank Control Warnings, trigger "2062_Warning_Data_BTCS_WARNING_WORD_05" bit 4
   2199: 'FIT420 5 PORT MBG FLOW HIGH', class Tank Control Warnings, trigger "2062_Warning_Data_BTCS_WARNING_WORD_05" bit 7
   2284: 'LT422 3 STARBOARD TANK LEVEL HIGH', class Tank Control Warnings, trigger "2062_Warning_Data_BTCS_WARNING_WORD_10" bit 12
   2198: 'FIT420 5 PORT MBG FLOW LOW', class Tank Control Warnings, trigger "2062_Warning_Data_BTCS_WARNING_WORD_05" bit 6
   2197: 'FIT419 4 STARBOARD MBG FLOW HIGH', class Tank Control Warnings, trigger "2062_Warning_Data_BTCS_WARNING_WORD_05" bit 5
   2283: 'LT422 3 PORT TANK LEVEL LOW', class Tank Control Warnings, trigger "2062_Warning_Data_BTCS_WARNING_WORD_10" bit 11
   2277: 'LT422 5 STARBOARD TANK LEVEL LOW', class Tank Control Warnings, trigger "2062_Warning_Data_BTCS_WARNING_WORD_10" bit 5
   2189: 'FIT417 4 STARBOARD TANK USD FLOW HIGH', class Tank Control Warnings, trigger "2062_Warning_Data_BTCS_WARNING_WORD_04" bit 13
   2188: 'FIT417 4 STARBOARD TANK USD FLOW LOW', class Tank Control Warnings, trigger "2062_Warning_Data_BTCS_WARNING_WORD_04" bit 12
   2276: 'LT422 5 STARBOARD TANK LEVEL HIGH', class Tank Control Warnings, trigger "2062_Warning_Data_BTCS_WARNING_WORD_10" bit 4
   2187: 'FIT418 4 PORT TANK USD FLOW HIGH', class Tank Control Warnings, trigger "2062_Warning_Data_BTCS_WARNING_WORD_04" bit 11
   2190: 'FIT418 5 PORT TANK USD FLOW LOW', class Tank Control Warnings, trigger "2062_Warning_Data_BTCS_WARNING_WORD_04" bit 14
   2192: 'FIT419 3 STARBOARD MBG FLOW LOW', class Tank Control Warnings, trigger "2062_Warning_Data_BTCS_WARNING_WORD_05" bit 0
   2280: 'LT422 2 STARBOARD TANK LEVEL HIGH', class Tank Control Warnings, trigger "2062_Warning_Data_BTCS_WARNING_WORD_10" bit 8
   2279: 'LT422 6 PORT TANK LEVEL LOW', class Tank Control Warnings, trigger "2062_Warning_Data_BTCS_WARNING_WORD_10" bit 7
   2278: 'LT422 6 PORT TANK LEVEL HIGH', class Tank Control Warnings, trigger "2062_Warning_Data_BTCS_WARNING_WORD_10" bit 6
   2191: 'FIT418 5 PORT TANK USD FLOW HIGH', class Tank Control Warnings, trigger "2062_Warning_Data_BTCS_WARNING_WORD_04" bit 15
   2167: 'FIT418 3 PORT TANK USD FLOW HIGH', class Tank Control Warnings, trigger "2062_Warning_Data_BTCS_WARNING_WORD_03" bit 7
   2061: 'PT415 RIO7 DECK IG PRESSURE HIGH HIGH', class Tank Control Alarms, trigger "2060_Alarm_Data_BTCS_ALARM_WORD_04" bit 13
   2062: '', class Tank Control Alarms, trigger "2060_Alarm_Data_BTCS_ALARM_WORD_04" bit 14
   2060: 'PT415 RIO7 DECK IG PRESSURE LOW LOW', class Tank Control Alarms, trigger "2060_Alarm_Data_BTCS_ALARM_WORD_04" bit 12
   2058: 'PT415 RIO6 DECK IG PRESSURE LOW LOW', class Tank Control Alarms, trigger "2060_Alarm_Data_BTCS_ALARM_WORD_04" bit 10
   2059: 'PT415 RIO6 DECK IG PRESSURE HGH HIGH', class Tank Control Alarms, trigger "2060_Alarm_Data_BTCS_ALARM_WORD_04" bit 11
   2063: '', class Tank Control Alarms, trigger "2060_Alarm_Data_BTCS_ALARM_WORD_04" bit 15
   2160: 'FIT418 1 FOR PEACK TANK USD FLOW LOW', class Tank Control Warnings, trigger "2062_Warning_Data_BTCS_WARNING_WORD_03" bit 0
   2161: 'FIT418 1 FOR PEACK TANK USD FLOW HIGH', class Tank Control Warnings, trigger "2062_Warning_Data_BTCS_WARNING_WORD_03" bit 1
